// TIA Portal project "SteviAutomation-ZadProg-DP_2" (V15.1)
// Przygotowanie logiki dla sterownika PLC Siemens S7-1200 zgodnie z opisem.

(* hardware
DEVICE "S7-1200 station_2"  S7-1200 Station
   slot 0: "Rack_0"  S7-1200 Rack  Rack  V1.0
   slot 1: "PLC_1"  CPU 1211C DC/DC/DC  6ES7 211-1AE40-0XB0  V4.2
DEVICE "PC-System_1"  SIMATIC PC station
   slot 0: "SIMATIC PC station"  Rail  SIMATIC PC-Station  V1.0
      slot 125: "Stationmanager"  Station_Manager  V6.0.4
   slot 1: "IE general_1"  IE General  IE_CP  V8.2.0
   slot 2: "HMI_RT_1"  WinCC RT Advanced  6AV2 104-0xxxx-xxxx  15.1.0.0
      slot 33792: "Host interface"  Host interface
*)

// ===== PLC "PLC_1"  CPU 1211C DC/DC/DC =====

VAR_GLOBAL   // PLC tag table "PLC_1"
   "Trigger_1" AT %I0.0 : Bool;   // State change trigger
   "Database_Full" AT %Q0.0 : Bool;   // Database is full
END_VAR

TYPE "SignalStatus"
   STRUCT
      sRecords : String;   // Single state change record
   END_STRUCT;
END_TYPE

TYPE "TimeStatic"
   STRUCT
      sYear : String;
      sMonth : String;
      sDay : String;
      sHour : String;
      sMinute : String;
      sSecond : String;
      sNanosecond : String;
   END_STRUCT;
END_TYPE

DATA_BLOCK "SaveRecord_DB"   // DB1
{ S7_Optimized_Access := 'TRUE' }
VERSION : 0.1
// stored: InstanceOfName SaveRecord_FB
"SaveRecord_FB"
BEGIN
END_DATA_BLOCK

DATA_BLOCK "DB_TriggerRecords"   // DB100
{ S7_Optimized_Access := 'TRUE' }
VERSION : 0.1
   VAR
      StateTable : Array[0..49] of "SignalStatus";   // Database containing state change records
      InitStateTable : Array[0..49] of "SignalStatus";   // Database containing state change records
      bAutoTrigger : Bool;   // Automode
      bAuxAutoManTrigger : Bool;
   END_VAR
BEGIN
END_DATA_BLOCK

FUNCTION_BLOCK "SaveRecord_FB"   // FB1, LAD
{ S7_Optimized_Access := 'TRUE' }
VERSION : 0.1
   VAR
      T_CONV : "T_CONV";   // Convert many to string
      iCurrent : Int;   // iteration
      bFirstScan : Bool;   // First scan
      usiRandomTtime : UDInt;   // Randomize time in automode
      Trigger_P : Bool;   // Rising edge - trigger
      Trigger_N : Bool;   // Falling edge - trigger
      Timer_1 : TON_TIME;   // AutoMode - time to switch on the trigger
      Timer_2 : TON_TIME;   // AutoMode - time to switch off the trigger
      tRandomTimeCurrent : Time;   // Timer_0 - Random time
      tRandomTimeCurrent_1 : Time;   // Timer_2 - Random time
      sState : String;   // State
      dtlLast : DTL;   // Time of last state
      dtlCurrent : DTL;   // Time of current state
      sTimeStamp : String;   // Timestamp
      sLastStatusTime : String;   // Time of last state
      tTimeLastState : Time;   // Time of last state
   END_VAR
   VAR RETAIN
      CTU_iCurrent : CTU_INT;   // CTU iCurrent
   END_VAR
   VAR
      bHiLo : Int;   // Trigger Tag HMI
      FB_Blink : "FB_Blink";   // Database full blinking
      bReset : Bool;   // Reset table with records
   END_VAR
   VAR_TEMP
      ret_val_RD_LOC_T : Word;
   END_VAR
   VAR_TEMP   // added for the SCL form of the ladder/FBD networks
      _w1 : Bool;
      _w2 : Bool;
      _w3 : Bool;
   END_VAR
BEGIN

REGION Network 1: State change trigger
   // Auto and manual mode
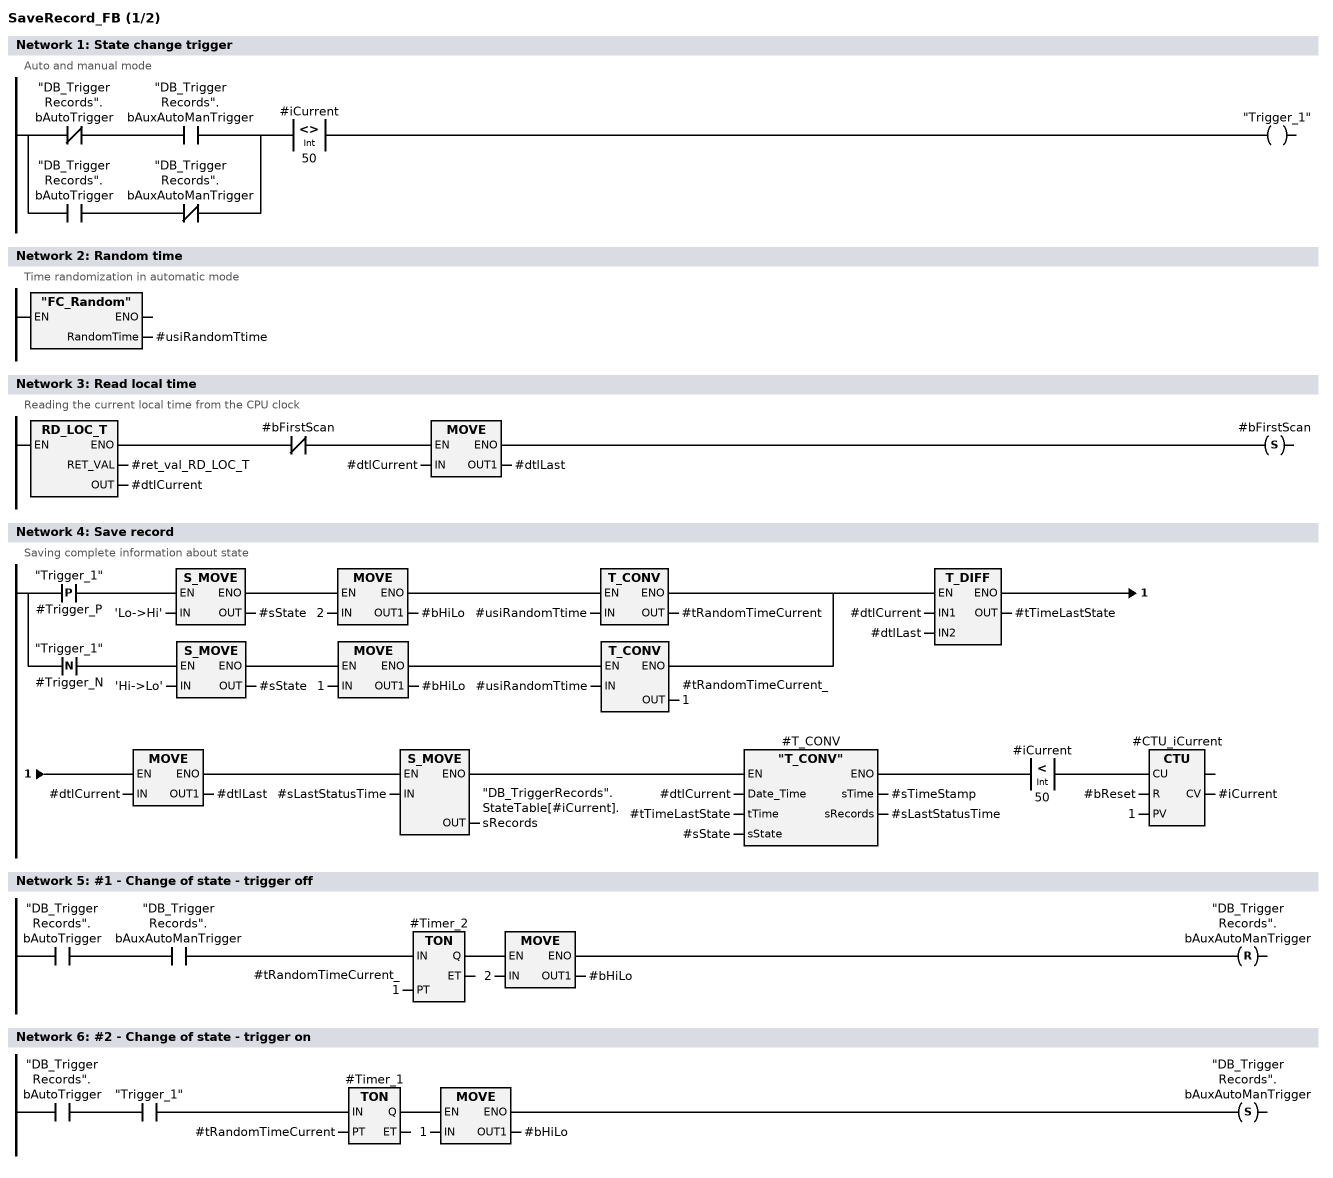
   RUNG wire#powerrail
      I_Contact( "DB_TriggerRecords".bAutoTrigger )
      Contact( "DB_TriggerRecords".bAuxAutoManTrigger )
      wire#w1
      { S7_Templates := "SrcType := Int" } NE_Contact(in1 := #iCurrent, in2 := 50)
      Coil( "Trigger_1" )
   END_RUNG
   RUNG wire#powerrail
      Contact( "DB_TriggerRecords".bAutoTrigger )
      I_Contact( "DB_TriggerRecords".bAuxAutoManTrigger )
   END_RUNG wire#w1
   // the same network as SCL:
   "Trigger_1" := ((NOT "DB_TriggerRecords".bAutoTrigger AND "DB_TriggerRecords".bAuxAutoManTrigger) OR ("DB_TriggerRecords".bAutoTrigger AND NOT "DB_TriggerRecords".bAuxAutoManTrigger)) AND (#iCurrent <> 50);
END_REGION

REGION Network 2: Random time
   // Time randomization in automatic mode
   RUNG wire#powerrail
      "FC_Random"(RandomTime => #usiRandomTtime)
   END_RUNG
   // the same network as SCL:
   "FC_Random"(RandomTime => #usiRandomTtime);
END_REGION

REGION Network 3: Read local time
   // Reading the current local time from the CPU clock
   // ENO of a box is taken as its EN; it also drops when the box reports an error
   #ret_val_RD_LOC_T := RD_LOC_T(OUT => #dtlCurrent);
   IF NOT #bFirstScan THEN
       #dtlLast := #dtlCurrent;
       #bFirstScan := TRUE;
   END_IF;
END_REGION

REGION Network 4: Save record
   // Saving complete information about state
   // ENO of a box is taken as its EN; it also drops when the box reports an error
   #_w1 := "Trigger_1" AND NOT #Trigger_P;   // rising edge of "Trigger_1"
   #Trigger_P := "Trigger_1";
   IF #_w1 THEN
       #sState := 'Lo->Hi';
       #bHiLo := 2;
       #tRandomTimeCurrent := T_CONV(IN := #usiRandomTtime);
   END_IF;
   #_w2 := NOT "Trigger_1" AND #Trigger_N;   // falling edge of "Trigger_1"
   #Trigger_N := "Trigger_1";
   IF #_w2 THEN
       #sState := 'Hi->Lo';
       #bHiLo := 1;
       #tRandomTimeCurrent_1 := T_CONV(IN := #usiRandomTtime);
   END_IF;
   IF #_w1 OR #_w2 THEN
       #tTimeLastState := T_DIFF(IN1 := #dtlCurrent, IN2 := #dtlLast);
       #dtlLast := #dtlCurrent;
       "DB_TriggerRecords".StateTable[#iCurrent].sRecords := #sLastStatusTime;
   END_IF;
   #T_CONV(EN := #_w1 OR #_w2,   // "T_CONV"
           Date_Time := #dtlCurrent,
           tTime := #tTimeLastState,
           sState := #sState,
           sTime => #sTimeStamp,
           sRecords => #sLastStatusTime,
           ENO => #_w3);
   #CTU_iCurrent(CU := #_w3 AND (#iCurrent < 50), R := #bReset, PV := 1, CV => #iCurrent);   // CTU
END_REGION

REGION Network 5: #1 - Change of state - trigger off
   #Timer_2(IN := "DB_TriggerRecords".bAutoTrigger AND "DB_TriggerRecords".bAuxAutoManTrigger,   // TON
            PT := #tRandomTimeCurrent_1);
   IF #Timer_2.Q THEN
       #bHiLo := 2;
       "DB_TriggerRecords".bAuxAutoManTrigger := FALSE;
   END_IF;
END_REGION

REGION Network 6: #2 - Change of state - trigger on
   #Timer_1(IN := "DB_TriggerRecords".bAutoTrigger AND "Trigger_1", PT := #tRandomTimeCurrent);   // TON
   IF #Timer_1.Q THEN
       #bHiLo := 1;
       "DB_TriggerRecords".bAuxAutoManTrigger := TRUE;
   END_IF;
END_REGION

REGION Network 7: Database full
   // In case of saving the last record - switching on the blinking with the [Database_full] output
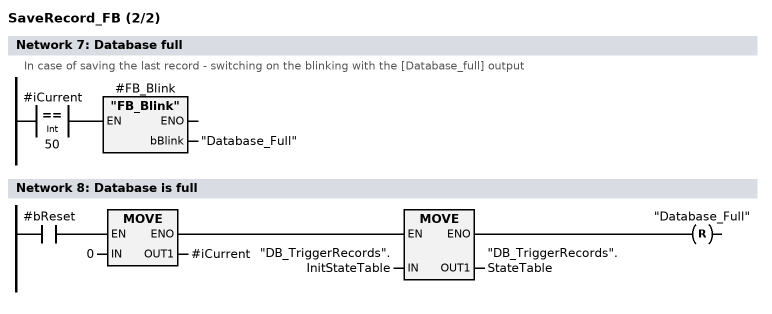
   RUNG wire#powerrail
      { S7_Templates := "SrcType := Int" } EQ_Contact(in1 := #iCurrent, in2 := 50)
      #FB_Blink(bBlink => "Database_Full")
   END_RUNG
   // the same network as SCL:
   IF #iCurrent = 50 THEN
       #FB_Blink(bBlink => "Database_Full");   // "FB_Blink"
   END_IF;
END_REGION

REGION Network 8: Database is full
   RUNG wire#powerrail
      Contact( #bReset )
      Move(in := 0, out1 => #iCurrent)
      Move(in := "DB_TriggerRecords".InitStateTable, out1 => "DB_TriggerRecords".StateTable)
      R_Coil( "Database_Full" )
   END_RUNG
   // the same network as SCL:
   IF #bReset THEN
       #iCurrent := 0;
       "DB_TriggerRecords".StateTable := "DB_TriggerRecords".InitStateTable;
       "Database_Full" := FALSE;
   END_IF;
END_REGION
END_FUNCTION_BLOCK

FUNCTION_BLOCK "FB_Blink"   // FB2, LAD
{ S7_Optimized_Access := 'TRUE' }
VERSION : 0.1
   VAR_OUTPUT
      bBlink : Bool;
   END_VAR
   VAR
      bBlinking : Bool;
      TON_Blink_off : TON_TIME;
      TON_Blink : TON_TIME;
   END_VAR
BEGIN

REGION Network 1: #bBlink
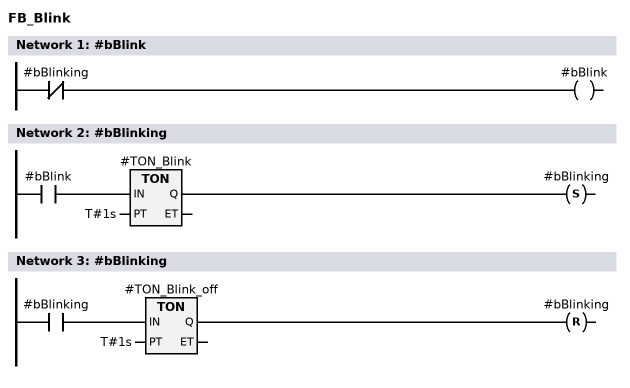
   RUNG wire#powerrail
      I_Contact( #bBlinking )
      Coil( #bBlink )
   END_RUNG
   // the same network as SCL:
   #bBlink := NOT #bBlinking;
END_REGION

REGION Network 2: #bBlinking
   #TON_Blink(IN := #bBlink, PT := T#1s);   // TON
   IF #TON_Blink.Q THEN #bBlinking := TRUE; END_IF;
END_REGION

REGION Network 3: #bBlinking
   #TON_Blink_off(IN := #bBlinking, PT := T#1s);   // TON
   IF #TON_Blink_off.Q THEN #bBlinking := FALSE; END_IF;
END_REGION
END_FUNCTION_BLOCK

FUNCTION_BLOCK "T_CONV"   // FB4, LAD
{ S7_Optimized_Access := 'TRUE' }
VERSION : 0.1
   VAR_INPUT
      Date_Time : DTL;   // Timestamp
      tTime : Time;   // Time of the previous state
      sState : String;   // State
   END_VAR
   VAR_OUTPUT
      sTime : String;   // Time of the previous state
      sRecords : String;   // Complete information about state
   END_VAR
   VAR
      sTimeStatic : "TimeStatic";
   END_VAR
   VAR_TEMP
      rRound : Real;   // Rounding of nanoseconds
      udiRounded : UDInt;   // Rounding of nanoseconds
      diTime : DInt;   // [auxiliary variable] Time of the previous state
      rTime : Real;   // [auxiliary variable] Time of the previous state
      sLastTime : String;   // Complete information about time
   END_VAR
   VAR_TEMP   // added for the SCL form of the ladder/FBD networks
      _w1 : Bool;
      _w2 : Bool;
   END_VAR
BEGIN

REGION Network 1: Initialize
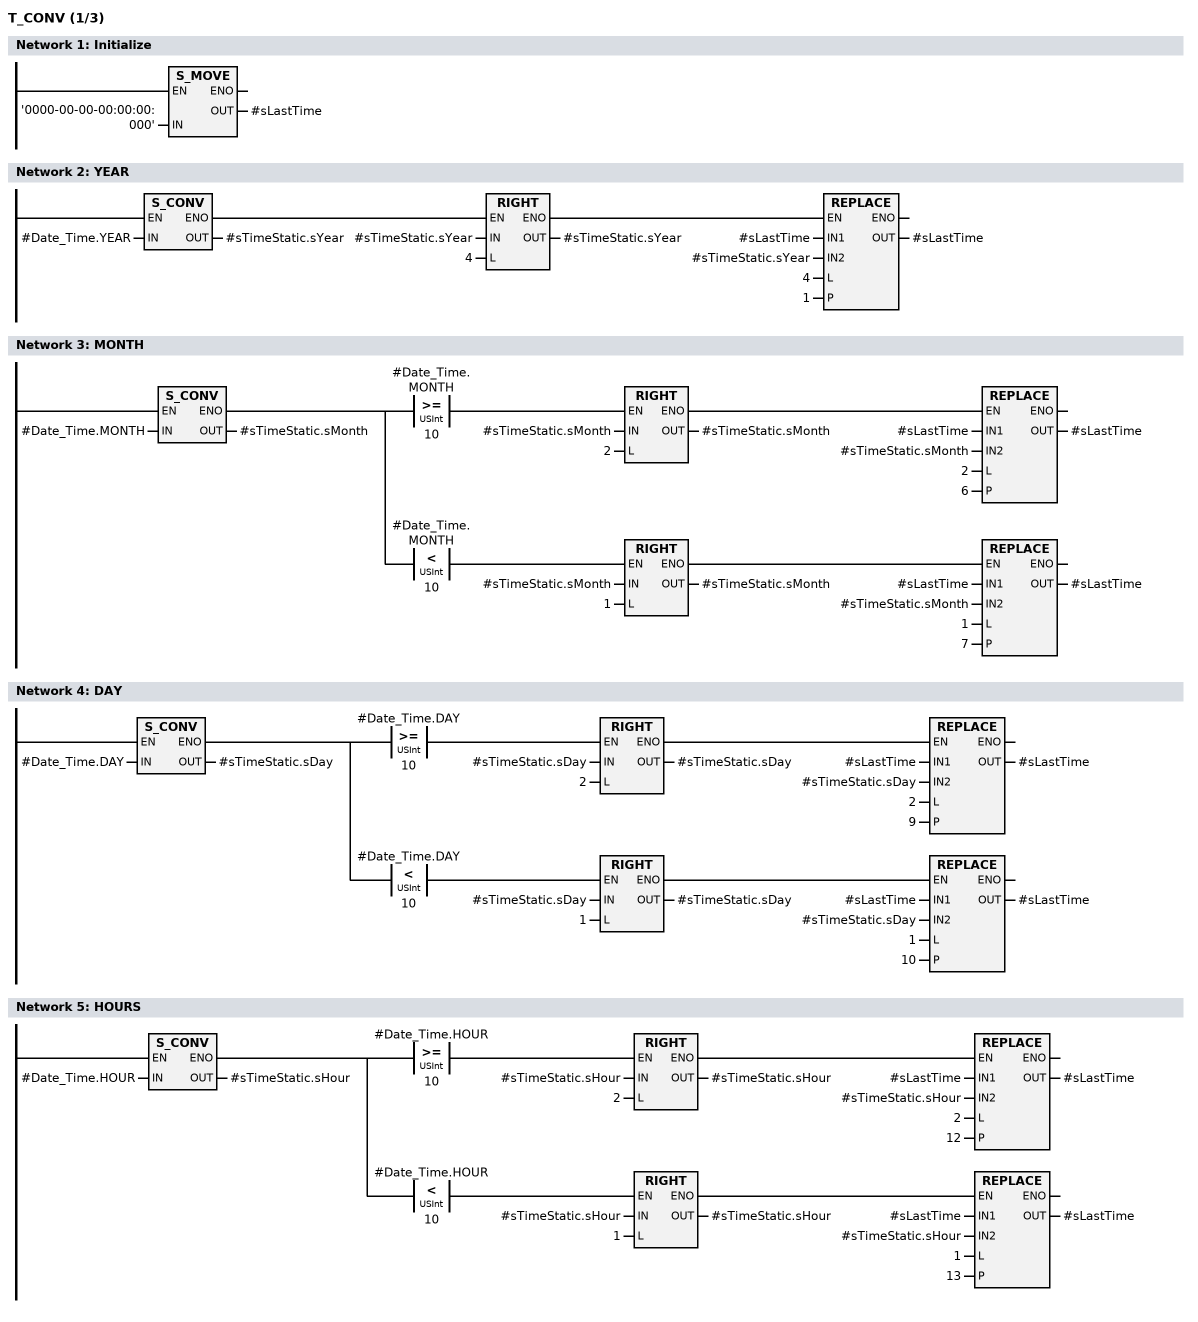
   RUNG wire#powerrail
      S_Move(in := '0000-00-00-00:00:00:000', out => #sLastTime)
   END_RUNG
   // the same network as SCL:
   #sLastTime := '0000-00-00-00:00:00:000';
END_REGION

REGION Network 2: YEAR
   #sTimeStatic.sYear := S_CONV(IN := #Date_Time.YEAR);
   #sTimeStatic.sYear := RIGHT(IN := #sTimeStatic.sYear, L := 4);
   #sLastTime := REPLACE(IN1 := #sLastTime, IN2 := #sTimeStatic.sYear, L := 4, P := 1);
END_REGION

REGION Network 3: MONTH
   #sTimeStatic.sMonth := S_CONV(IN := #Date_Time.MONTH);
   IF #Date_Time.MONTH >= 10 THEN
       #sTimeStatic.sMonth := RIGHT(IN := #sTimeStatic.sMonth, L := 2);
       #sLastTime := REPLACE(IN1 := #sLastTime, IN2 := #sTimeStatic.sMonth, L := 2, P := 6);
   END_IF;
   IF #Date_Time.MONTH < 10 THEN
       #sTimeStatic.sMonth := RIGHT(IN := #sTimeStatic.sMonth, L := 1);
       #sLastTime := REPLACE(IN1 := #sLastTime, IN2 := #sTimeStatic.sMonth, L := 1, P := 7);
   END_IF;
END_REGION

REGION Network 4: DAY
   #sTimeStatic.sDay := S_CONV(IN := #Date_Time.DAY);
   IF #Date_Time.DAY >= 10 THEN
       #sTimeStatic.sDay := RIGHT(IN := #sTimeStatic.sDay, L := 2);
       #sLastTime := REPLACE(IN1 := #sLastTime, IN2 := #sTimeStatic.sDay, L := 2, P := 9);
   END_IF;
   IF #Date_Time.DAY < 10 THEN
       #sTimeStatic.sDay := RIGHT(IN := #sTimeStatic.sDay, L := 1);
       #sLastTime := REPLACE(IN1 := #sLastTime, IN2 := #sTimeStatic.sDay, L := 1, P := 10);
   END_IF;
END_REGION

REGION Network 5: HOURS
   #sTimeStatic.sHour := S_CONV(IN := #Date_Time.HOUR);
   IF #Date_Time.HOUR >= 10 THEN
       #sTimeStatic.sHour := RIGHT(IN := #sTimeStatic.sHour, L := 2);
       #sLastTime := REPLACE(IN1 := #sLastTime, IN2 := #sTimeStatic.sHour, L := 2, P := 12);
   END_IF;
   IF #Date_Time.HOUR < 10 THEN
       #sTimeStatic.sHour := RIGHT(IN := #sTimeStatic.sHour, L := 1);
       #sLastTime := REPLACE(IN1 := #sLastTime, IN2 := #sTimeStatic.sHour, L := 1, P := 13);
   END_IF;
END_REGION

REGION Network 6: MINUTES
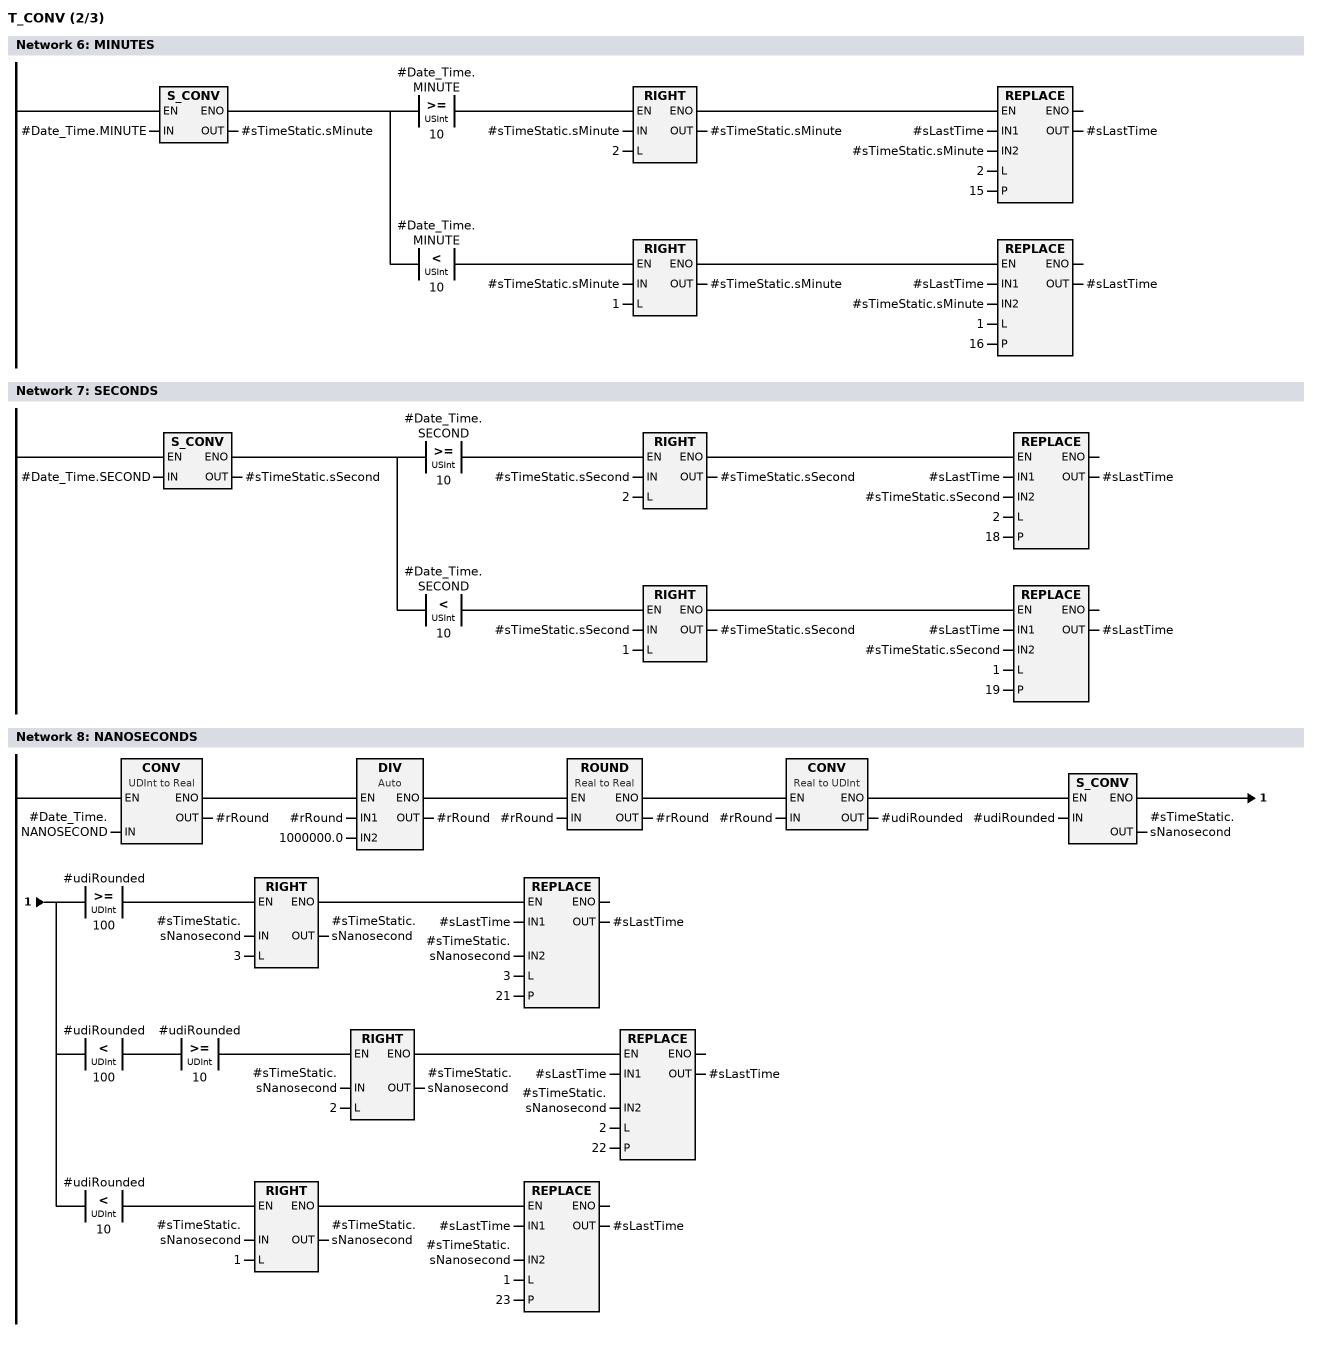
   #sTimeStatic.sMinute := S_CONV(IN := #Date_Time.MINUTE);
   IF #Date_Time.MINUTE >= 10 THEN
       #sTimeStatic.sMinute := RIGHT(IN := #sTimeStatic.sMinute, L := 2);
       #sLastTime := REPLACE(IN1 := #sLastTime, IN2 := #sTimeStatic.sMinute, L := 2, P := 15);
   END_IF;
   IF #Date_Time.MINUTE < 10 THEN
       #sTimeStatic.sMinute := RIGHT(IN := #sTimeStatic.sMinute, L := 1);
       #sLastTime := REPLACE(IN1 := #sLastTime, IN2 := #sTimeStatic.sMinute, L := 1, P := 16);
   END_IF;
END_REGION

REGION Network 7: SECONDS
   #sTimeStatic.sSecond := S_CONV(IN := #Date_Time.SECOND);
   IF #Date_Time.SECOND >= 10 THEN
       #sTimeStatic.sSecond := RIGHT(IN := #sTimeStatic.sSecond, L := 2);
       #sLastTime := REPLACE(IN1 := #sLastTime, IN2 := #sTimeStatic.sSecond, L := 2, P := 18);
   END_IF;
   IF #Date_Time.SECOND < 10 THEN
       #sTimeStatic.sSecond := RIGHT(IN := #sTimeStatic.sSecond, L := 1);
       #sLastTime := REPLACE(IN1 := #sLastTime, IN2 := #sTimeStatic.sSecond, L := 1, P := 19);
   END_IF;
END_REGION

REGION Network 8: NANOSECONDS
   #rRound := UDINT_TO_REAL(#Date_Time.NANOSECOND);
   #rRound := #rRound / 1000000.0;
   #rRound := ROUND(#rRound);
   #udiRounded := REAL_TO_UDINT(#rRound);
   #sTimeStatic.sNanosecond := S_CONV(IN := #udiRounded);
   IF #udiRounded >= 100 THEN
       #sTimeStatic.sNanosecond := RIGHT(IN := #sTimeStatic.sNanosecond, L := 3);
       #sLastTime := REPLACE(IN1 := #sLastTime, IN2 := #sTimeStatic.sNanosecond, L := 3, P := 21);
   END_IF;
   IF (#udiRounded < 100) AND (#udiRounded >= 10) THEN
       #sTimeStatic.sNanosecond := RIGHT(IN := #sTimeStatic.sNanosecond, L := 2);
       #sLastTime := REPLACE(IN1 := #sLastTime, IN2 := #sTimeStatic.sNanosecond, L := 2, P := 22);
   END_IF;
   IF #udiRounded < 10 THEN
       #sTimeStatic.sNanosecond := RIGHT(IN := #sTimeStatic.sNanosecond, L := 1);
       #sLastTime := REPLACE(IN1 := #sLastTime, IN2 := #sTimeStatic.sNanosecond, L := 1, P := 23);
   END_IF;
END_REGION

REGION Network 9: #1 - Time of the previous state
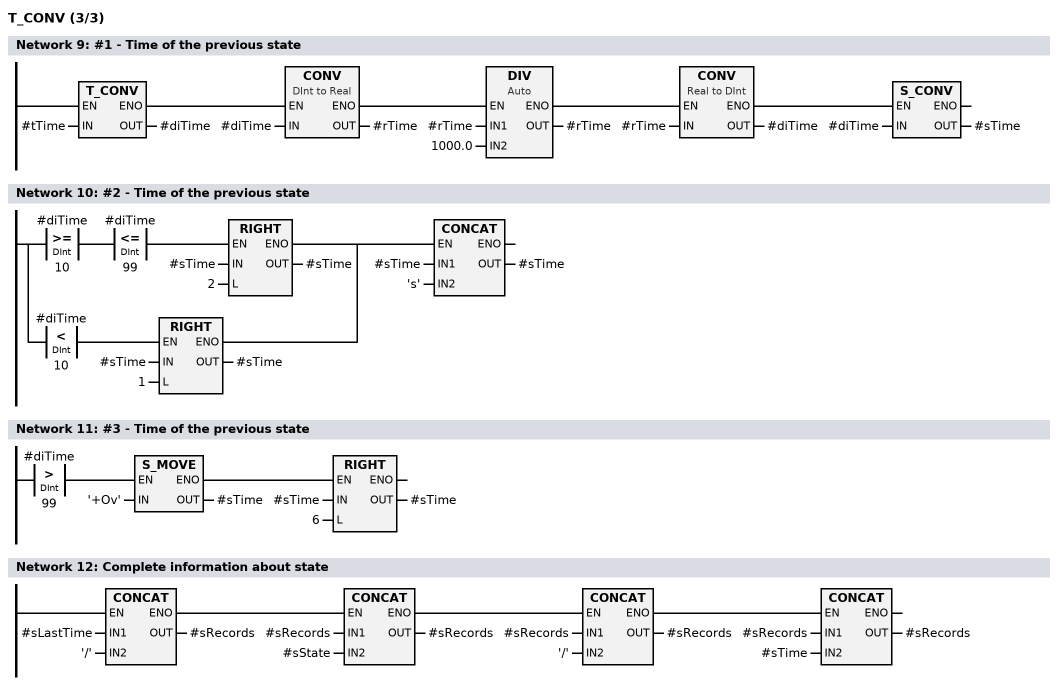
   // ENO of a box is taken as its EN; it also drops when the box reports an error
   #diTime := T_CONV(IN := #tTime);
   #rTime := DINT_TO_REAL(#diTime);
   #rTime := #rTime / 1000.0;
   #diTime := REAL_TO_DINT(#rTime);
   #sTime := S_CONV(IN := #diTime);
END_REGION

REGION Network 10: #2 - Time of the previous state
   #_w1 := (#diTime >= 10) AND (#diTime <= 99);
   IF #_w1 THEN #sTime := RIGHT(IN := #sTime, L := 2); END_IF;
   #_w2 := #diTime < 10;
   IF #_w2 THEN #sTime := RIGHT(IN := #sTime, L := 1); END_IF;
   IF #_w1 OR #_w2 THEN #sTime := CONCAT(IN1 := #sTime, IN2 := 's'); END_IF;
END_REGION

REGION Network 11: #3 - Time of the previous state
   IF #diTime > 99 THEN
       #sTime := '+Ov';
       #sTime := RIGHT(IN := #sTime, L := 6);
   END_IF;
END_REGION

REGION Network 12: Complete information about state
   #sRecords := CONCAT(IN1 := #sLastTime, IN2 := '/');
   #sRecords := CONCAT(IN1 := #sRecords, IN2 := #sState);
   #sRecords := CONCAT(IN1 := #sRecords, IN2 := '/');
   #sRecords := CONCAT(IN1 := #sRecords, IN2 := #sTime);
END_REGION
END_FUNCTION_BLOCK

FUNCTION "FC_Random" : Void   // FC3, LAD
{ S7_Optimized_Access := 'TRUE' }
VERSION : 0.1
   VAR_OUTPUT
      RandomTime : UDInt;
   END_VAR
   VAR_TEMP
      time_Ret_Val : Int;
      PLC_System_Time : DTL;
   END_VAR
BEGIN

REGION Network 1: Draw from a range 0 - 120000 (Udint)
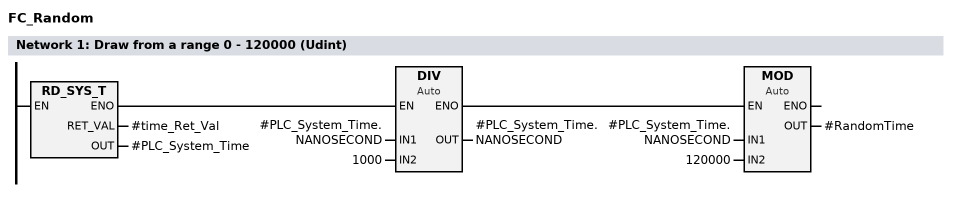
   // ENO of a box is taken as its EN; it also drops when the box reports an error
   #time_Ret_Val := RD_SYS_T(OUT => #PLC_System_Time);
   #PLC_System_Time.NANOSECOND := #PLC_System_Time.NANOSECOND / 1000;
   #RandomTime := #PLC_System_Time.NANOSECOND MOD 120000;
END_REGION
END_FUNCTION

ORGANIZATION_BLOCK "Main"   // OB1, LAD, ProgramCycle
TITLE = "Main Program Sweep (Cycle)"
{ S7_Optimized_Access := 'TRUE' }
VERSION : 0.1
   VAR_INPUT
      Initial_Call : Bool;   // Initial call of this OB
      Remanence : Bool;   // =True, if remanent data are available
   END_VAR
BEGIN

REGION Network 1: Saving records to table
   // Main logic responsible for checking the signal Trigger_1 (% I0.0). Each rising and falling edge is saving in the database with the current time stamp and the time of the previous state. The database contains 50 records.
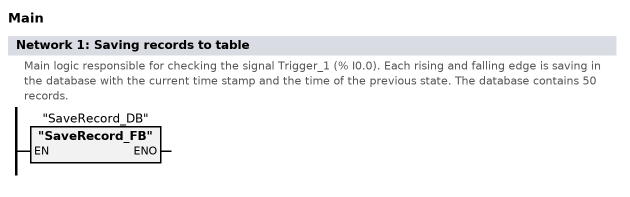
   RUNG wire#powerrail
      "SaveRecord_DB"()
   END_RUNG
   // the same network as SCL:
   "SaveRecord_DB"();   // "SaveRecord_FB"
END_REGION
END_ORGANIZATION_BLOCK

(* ===== HMI "HMI_RT_1" =====
system functions are stored by id; their names below are inferred from use
connection "HMI_Connection_1": ETHERNET, S7_1200_OMS

HMI tags "Default tag table"
   "Database_Full" : Bool = PLC Database_Full AT %Q0.0, 1 s
   "SaveRecord_DB_iCurrent" : Int = PLC SaveRecord_DB.iCurrent, 1 s
   "SaveRecord_DB_bReset" : Bool = PLC SaveRecord_DB.bReset, 1 s
   "Trigger_1" : Bool = PLC Trigger_1 AT %I0.0, 1 s

HMI tags "Events"
   "Record" : String[254] = PLC SaveRecord_DB.sLastStatusTime AT %DB1.DBW0, 1 s
   "HiLo" : Int = PLC SaveRecord_DB.bHiLo AT %DB1.DBX0.0, 1 s
   "TriggerButton" : Bool = PLC DB_TriggerRecords.bAuxAutoManTrigger AT %DB1.DBX0.0, 1 s
   "AutoMan" : Bool = PLC DB_TriggerRecords.bAutoTrigger AT %DB1.DBX0.0, 1 s

discrete alarms
   1: ')', class Status, trigger "HiLo" bit 1

screen "Screen_1" 1024x768
   Button "Button_1" at 820,157 size 153x78; TextOff 'Change State'
      on Click: InvertBit("TriggerButton")
      Appearance <- "Trigger_1"
      ObjectEnable <- "SaveRecord_DB_iCurrent"
   AlarmView "Alarm view_1" at 78,73 size 704x647; ColumnTextNumber 'No. / Nr / N.º.'; ColumnTextTime 'Time / Czas / Hora'; ColumnTextDate 'Data / Fecha'; ColumnTextAlarmText 'Records / Tekst / Texto'
   Rectangle "Rectangle_1" at 99,20 size 665x50
      Visibility <- "Database_Full"
   TextField "Text field_1" at 322,29 size 172x34; Text 'Database full'
      Visibility <- "Database_Full"
   Button "Button_2" at 820,252 size 153x78; TextOff 'Reset'
      on Press: function_b14e0dd5("SaveRecord_DB_bReset", 0)
   DateTimeField "Date/time field_1" at 792,29 size 212x31
   Switch "Switch_1" at 841,75 size 120x65; CaptionText 'Manual / Auto'; TextOff 'OFF'; TextOn 'ON'
      Appearance <- "AutoMan"
      ProcessValue <- "AutoMan"
      on Change: InvertBit("AutoMan")
      ObjectEnable <- "SaveRecord_DB_iCurrent"
*)